REGION Network 43
   RUNG wire#powerrail
      Contact( "DB92".Static_1 )
      { S7_GenerateENO := "TRUE" } Move(in := 1, out1 => "DB46".Static_19)
      wire#w1
      Coil( "Tag_6" )
   END_RUNG
   RUNG wire#powerrail
      I_Contact( "DB92".Static_1 )
      { S7_GenerateENO := "TRUE" } Move(in := 2, out1 => "DB46".Static_19)
   END_RUNG wire#w1
   // the same network as SCL:
   // ENO of a box is taken as its EN; it also drops when the box reports an error
   IF "DB92".Static_1 THEN "DB46".Static_19 := 1; END_IF;
   IF NOT "DB92".Static_1 THEN "DB46".Static_19 := 2; END_IF;
   "Tag_6" := "DB92".Static_1 OR NOT "DB92".Static_1;
END_REGION

REGION Network 44
   RUNG wire#powerrail
      Contact( "DB92".Static_2 )
      { S7_GenerateENO := "TRUE" } Move(in := 1, out1 => "DB46".Static_20)
      wire#w1
      Coil( "Tag_6" )
   END_RUNG
   RUNG wire#powerrail
      I_Contact( "DB92".Static_2 )
      { S7_GenerateENO := "TRUE" } Move(in := 2, out1 => "DB46".Static_20)
   END_RUNG wire#w1
   // the same network as SCL:
   // ENO of a box is taken as its EN; it also drops when the box reports an error
   IF "DB92".Static_2 THEN "DB46".Static_20 := 1; END_IF;
   IF NOT "DB92".Static_2 THEN "DB46".Static_20 := 2; END_IF;
   "Tag_6" := "DB92".Static_2 OR NOT "DB92".Static_2;
END_REGION

REGION Network 45
   RUNG wire#powerrail
      Contact( "DB21".Static_52 )
      { S7_GenerateENO := "TRUE" } Move(in := 1, out1 => "DB46".Static_23)
      wire#w1
      Coil( "Tag_6" )
   END_RUNG
   RUNG wire#powerrail
      I_Contact( "DB21".Static_52 )
      { S7_GenerateENO := "TRUE" } Move(in := 2, out1 => "DB46".Static_23)
   END_RUNG wire#w1
   // the same network as SCL:
   // ENO of a box is taken as its EN; it also drops when the box reports an error
   IF "DB21".Static_52 THEN "DB46".Static_23 := 1; END_IF;
   IF NOT "DB21".Static_52 THEN "DB46".Static_23 := 2; END_IF;
   "Tag_6" := "DB21".Static_52 OR NOT "DB21".Static_52;
END_REGION

REGION Network 46
   RUNG wire#powerrail
      Contact( "DB21".Static_53 )
      { S7_GenerateENO := "TRUE" } Move(in := 1, out1 => "DB46".Static_24)
      wire#w1
      Coil( "Tag_6" )
   END_RUNG
   RUNG wire#powerrail
      I_Contact( "DB21".Static_53 )
      { S7_GenerateENO := "TRUE" } Move(in := 2, out1 => "DB46".Static_24)
   END_RUNG wire#w1
   // the same network as SCL:
   // ENO of a box is taken as its EN; it also drops when the box reports an error
   IF "DB21".Static_53 THEN "DB46".Static_24 := 1; END_IF;
   IF NOT "DB21".Static_53 THEN "DB46".Static_24 := 2; END_IF;
   "Tag_6" := "DB21".Static_53 OR NOT "DB21".Static_53;
END_REGION

REGION Network 47
   RUNG wire#powerrail
      Contact( "DB135".Static_18 )
      { S7_GenerateENO := "TRUE" } Move(in := 0, out1 => "DB135".Static_0)
      wire#w1
      Coil( "Tag_6" )
   END_RUNG
   RUNG wire#powerrail
      I_Contact( "DB135".Static_18 )
      Contact( "DB88".Static_12 )
      { S7_GenerateENO := "TRUE" } Move(in := 1, out1 => "DB135".Static_0)
   END_RUNG wire#w1
   RUNG wire#powerrail
      I_Contact( "DB135".Static_18 )
      I_Contact( "DB88".Static_12 )
      { S7_GenerateENO := "TRUE" } Move(in := 2, out1 => "DB135".Static_0)
   END_RUNG wire#w1
   // the same network as SCL:
   // ENO of a box is taken as its EN; it also drops when the box reports an error
   IF "DB135".Static_18 THEN "DB135".Static_0 := 0; END_IF;
   #_w1 := NOT "DB135".Static_18 AND "DB88".Static_12;
   IF #_w1 THEN "DB135".Static_0 := 1; END_IF;
   #_w2 := NOT "DB135".Static_18 AND NOT "DB88".Static_12;
   IF #_w2 THEN "DB135".Static_0 := 2; END_IF;
   "Tag_6" := "DB135".Static_18 OR #_w1 OR #_w2;
END_REGION

REGION Network 48
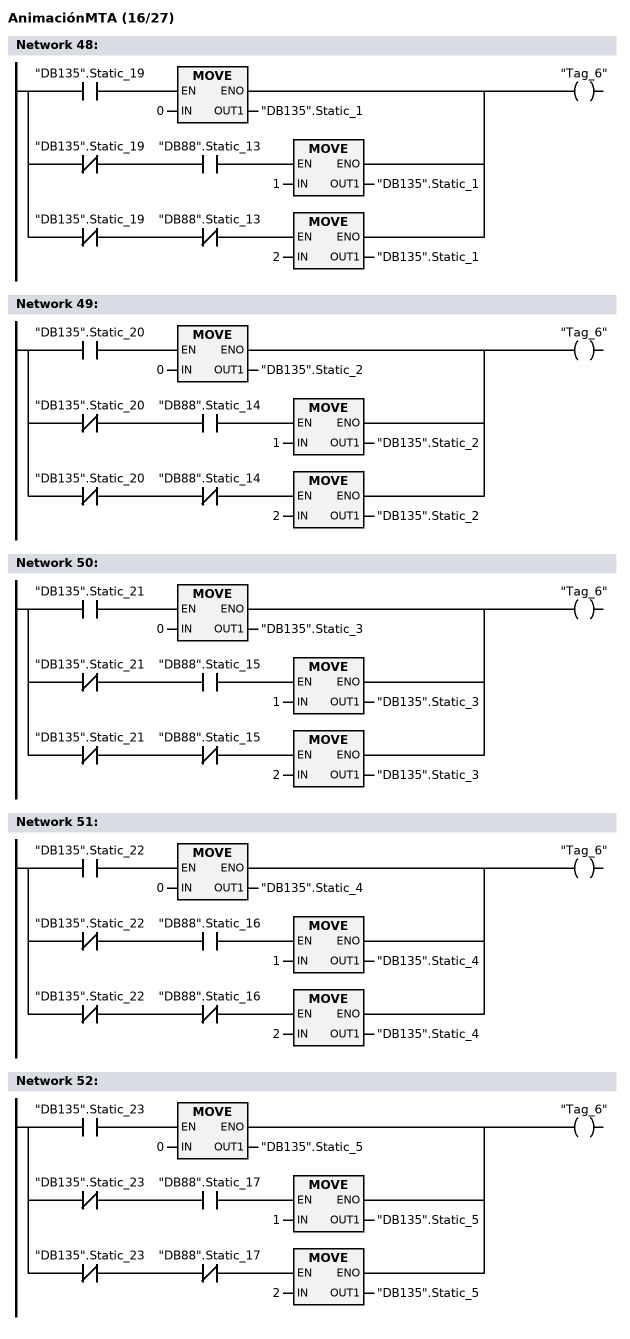
   RUNG wire#powerrail
      Contact( "DB135".Static_19 )
      { S7_GenerateENO := "TRUE" } Move(in := 0, out1 => "DB135".Static_1)
      wire#w1
      Coil( "Tag_6" )
   END_RUNG
   RUNG wire#powerrail
      I_Contact( "DB135".Static_19 )
      Contact( "DB88".Static_13 )
      { S7_GenerateENO := "TRUE" } Move(in := 1, out1 => "DB135".Static_1)
   END_RUNG wire#w1
   RUNG wire#powerrail
      I_Contact( "DB135".Static_19 )
      I_Contact( "DB88".Static_13 )
      { S7_GenerateENO := "TRUE" } Move(in := 2, out1 => "DB135".Static_1)
   END_RUNG wire#w1
   // the same network as SCL:
   // ENO of a box is taken as its EN; it also drops when the box reports an error
   IF "DB135".Static_19 THEN "DB135".Static_1 := 0; END_IF;
   #_w1 := NOT "DB135".Static_19 AND "DB88".Static_13;
   IF #_w1 THEN "DB135".Static_1 := 1; END_IF;
   #_w2 := NOT "DB135".Static_19 AND NOT "DB88".Static_13;
   IF #_w2 THEN "DB135".Static_1 := 2; END_IF;
   "Tag_6" := "DB135".Static_19 OR #_w1 OR #_w2;
END_REGION

REGION Network 49
   RUNG wire#powerrail
      Contact( "DB135".Static_20 )
      { S7_GenerateENO := "TRUE" } Move(in := 0, out1 => "DB135".Static_2)
      wire#w1
      Coil( "Tag_6" )
   END_RUNG
   RUNG wire#powerrail
      I_Contact( "DB135".Static_20 )
      Contact( "DB88".Static_14 )
      { S7_GenerateENO := "TRUE" } Move(in := 1, out1 => "DB135".Static_2)
   END_RUNG wire#w1
   RUNG wire#powerrail
      I_Contact( "DB135".Static_20 )
      I_Contact( "DB88".Static_14 )
      { S7_GenerateENO := "TRUE" } Move(in := 2, out1 => "DB135".Static_2)
   END_RUNG wire#w1
   // the same network as SCL:
   // ENO of a box is taken as its EN; it also drops when the box reports an error
   IF "DB135".Static_20 THEN "DB135".Static_2 := 0; END_IF;
   #_w1 := NOT "DB135".Static_20 AND "DB88".Static_14;
   IF #_w1 THEN "DB135".Static_2 := 1; END_IF;
   #_w2 := NOT "DB135".Static_20 AND NOT "DB88".Static_14;
   IF #_w2 THEN "DB135".Static_2 := 2; END_IF;
   "Tag_6" := "DB135".Static_20 OR #_w1 OR #_w2;
END_REGION

REGION Network 50
   RUNG wire#powerrail
      Contact( "DB135".Static_21 )
      { S7_GenerateENO := "TRUE" } Move(in := 0, out1 => "DB135".Static_3)
      wire#w1
      Coil( "Tag_6" )
   END_RUNG
   RUNG wire#powerrail
      I_Contact( "DB135".Static_21 )
      Contact( "DB88".Static_15 )
      { S7_GenerateENO := "TRUE" } Move(in := 1, out1 => "DB135".Static_3)
   END_RUNG wire#w1
   RUNG wire#powerrail
      I_Contact( "DB135".Static_21 )
      I_Contact( "DB88".Static_15 )
      { S7_GenerateENO := "TRUE" } Move(in := 2, out1 => "DB135".Static_3)
   END_RUNG wire#w1
   // the same network as SCL:
   // ENO of a box is taken as its EN; it also drops when the box reports an error
   IF "DB135".Static_21 THEN "DB135".Static_3 := 0; END_IF;
   #_w1 := NOT "DB135".Static_21 AND "DB88".Static_15;
   IF #_w1 THEN "DB135".Static_3 := 1; END_IF;
   #_w2 := NOT "DB135".Static_21 AND NOT "DB88".Static_15;
   IF #_w2 THEN "DB135".Static_3 := 2; END_IF;
   "Tag_6" := "DB135".Static_21 OR #_w1 OR #_w2;
END_REGION

REGION Network 51
   RUNG wire#powerrail
      Contact( "DB135".Static_22 )
      { S7_GenerateENO := "TRUE" } Move(in := 0, out1 => "DB135".Static_4)
      wire#w1
      Coil( "Tag_6" )
   END_RUNG
   RUNG wire#powerrail
      I_Contact( "DB135".Static_22 )
      Contact( "DB88".Static_16 )
      { S7_GenerateENO := "TRUE" } Move(in := 1, out1 => "DB135".Static_4)
   END_RUNG wire#w1
   RUNG wire#powerrail
      I_Contact( "DB135".Static_22 )
      I_Contact( "DB88".Static_16 )
      { S7_GenerateENO := "TRUE" } Move(in := 2, out1 => "DB135".Static_4)
   END_RUNG wire#w1
   // the same network as SCL:
   // ENO of a box is taken as its EN; it also drops when the box reports an error
   IF "DB135".Static_22 THEN "DB135".Static_4 := 0; END_IF;
   #_w1 := NOT "DB135".Static_22 AND "DB88".Static_16;
   IF #_w1 THEN "DB135".Static_4 := 1; END_IF;
   #_w2 := NOT "DB135".Static_22 AND NOT "DB88".Static_16;
   IF #_w2 THEN "DB135".Static_4 := 2; END_IF;
   "Tag_6" := "DB135".Static_22 OR #_w1 OR #_w2;
END_REGION

REGION Network 52
   RUNG wire#powerrail
      Contact( "DB135".Static_23 )
      { S7_GenerateENO := "TRUE" } Move(in := 0, out1 => "DB135".Static_5)
      wire#w1
      Coil( "Tag_6" )
   END_RUNG
   RUNG wire#powerrail
      I_Contact( "DB135".Static_23 )
      Contact( "DB88".Static_17 )
      { S7_GenerateENO := "TRUE" } Move(in := 1, out1 => "DB135".Static_5)
   END_RUNG wire#w1
   RUNG wire#powerrail
      I_Contact( "DB135".Static_23 )
      I_Contact( "DB88".Static_17 )
      { S7_GenerateENO := "TRUE" } Move(in := 2, out1 => "DB135".Static_5)
   END_RUNG wire#w1
   // the same network as SCL:
   // ENO of a box is taken as its EN; it also drops when the box reports an error
   IF "DB135".Static_23 THEN "DB135".Static_5 := 0; END_IF;
   #_w1 := NOT "DB135".Static_23 AND "DB88".Static_17;
   IF #_w1 THEN "DB135".Static_5 := 1; END_IF;
   #_w2 := NOT "DB135".Static_23 AND NOT "DB88".Static_17;
   IF #_w2 THEN "DB135".Static_5 := 2; END_IF;
   "Tag_6" := "DB135".Static_23 OR #_w1 OR #_w2;
END_REGION

REGION Network 53
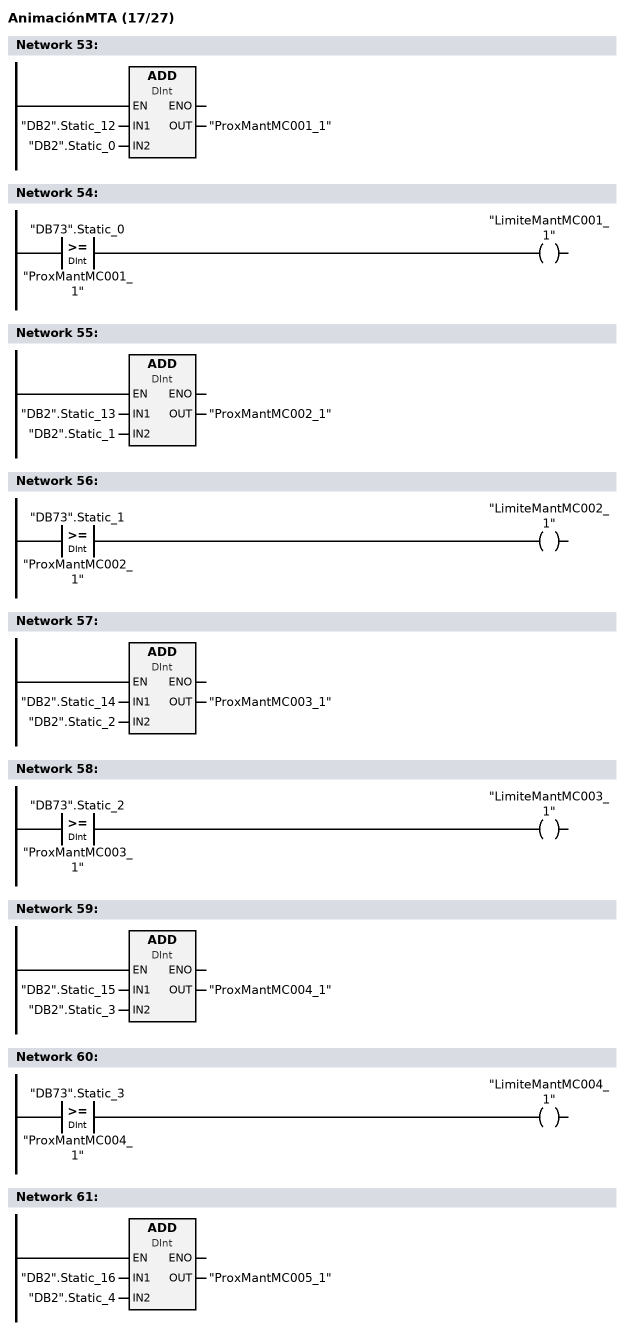
   RUNG wire#powerrail
      { S7_Templates := "SrcType := DInt"; S7_GenerateENO := "TRUE" } Add(in1 := "DB2".Static_12, in2 := "DB2".Static_0, out => "ProxMantMC001_1")
   END_RUNG
   // the same network as SCL:
   "ProxMantMC001_1" := "DB2".Static_12 + "DB2".Static_0;
END_REGION

REGION Network 54
   RUNG wire#powerrail
      { S7_Templates := "SrcType := DInt" } GE_Contact(in1 := "DB73".Static_0, in2 := "ProxMantMC001_1")
      Coil( "LimiteMantMC001_1" )
   END_RUNG
   // the same network as SCL:
   "LimiteMantMC001_1" := "DB73".Static_0 >= "ProxMantMC001_1";
END_REGION

REGION Network 55
   RUNG wire#powerrail
      { S7_Templates := "SrcType := DInt"; S7_GenerateENO := "TRUE" } Add(in1 := "DB2".Static_13, in2 := "DB2".Static_1, out => "ProxMantMC002_1")
   END_RUNG
   // the same network as SCL:
   "ProxMantMC002_1" := "DB2".Static_13 + "DB2".Static_1;
END_REGION

REGION Network 56
   RUNG wire#powerrail
      { S7_Templates := "SrcType := DInt" } GE_Contact(in1 := "DB73".Static_1, in2 := "ProxMantMC002_1")
      Coil( "LimiteMantMC002_1" )
   END_RUNG
   // the same network as SCL:
   "LimiteMantMC002_1" := "DB73".Static_1 >= "ProxMantMC002_1";
END_REGION

REGION Network 57
   RUNG wire#powerrail
      { S7_Templates := "SrcType := DInt"; S7_GenerateENO := "TRUE" } Add(in1 := "DB2".Static_14, in2 := "DB2".Static_2, out => "ProxMantMC003_1")
   END_RUNG
   // the same network as SCL:
   "ProxMantMC003_1" := "DB2".Static_14 + "DB2".Static_2;
END_REGION

REGION Network 58
   RUNG wire#powerrail
      { S7_Templates := "SrcType := DInt" } GE_Contact(in1 := "DB73".Static_2, in2 := "ProxMantMC003_1")
      Coil( "LimiteMantMC003_1" )
   END_RUNG
   // the same network as SCL:
   "LimiteMantMC003_1" := "DB73".Static_2 >= "ProxMantMC003_1";
END_REGION

REGION Network 59
   RUNG wire#powerrail
      { S7_Templates := "SrcType := DInt"; S7_GenerateENO := "TRUE" } Add(in1 := "DB2".Static_15, in2 := "DB2".Static_3, out => "ProxMantMC004_1")
   END_RUNG
   // the same network as SCL:
   "ProxMantMC004_1" := "DB2".Static_15 + "DB2".Static_3;
END_REGION

REGION Network 60
   RUNG wire#powerrail
      { S7_Templates := "SrcType := DInt" } GE_Contact(in1 := "DB73".Static_3, in2 := "ProxMantMC004_1")
      Coil( "LimiteMantMC004_1" )
   END_RUNG
   // the same network as SCL:
   "LimiteMantMC004_1" := "DB73".Static_3 >= "ProxMantMC004_1";
END_REGION

REGION Network 61
   RUNG wire#powerrail
      { S7_Templates := "SrcType := DInt"; S7_GenerateENO := "TRUE" } Add(in1 := "DB2".Static_16, in2 := "DB2".Static_4, out => "ProxMantMC005_1")
   END_RUNG
   // the same network as SCL:
   "ProxMantMC005_1" := "DB2".Static_16 + "DB2".Static_4;
END_REGION

REGION Network 62
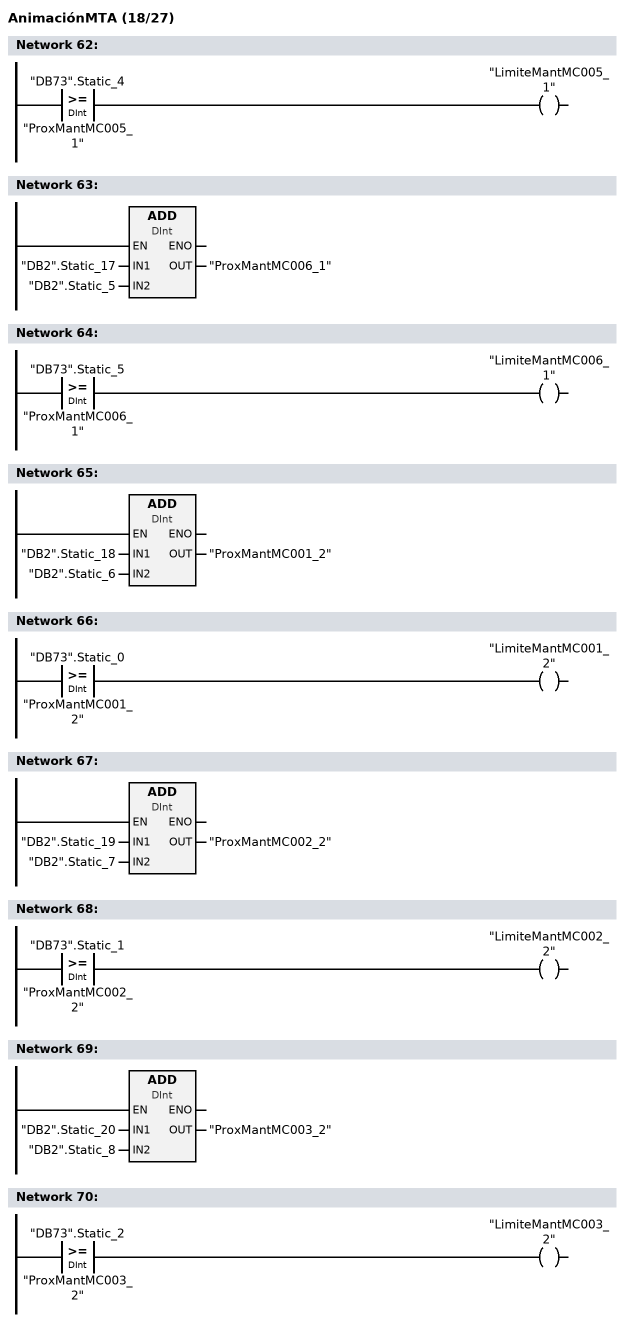
   RUNG wire#powerrail
      { S7_Templates := "SrcType := DInt" } GE_Contact(in1 := "DB73".Static_4, in2 := "ProxMantMC005_1")
      Coil( "LimiteMantMC005_1" )
   END_RUNG
   // the same network as SCL:
   "LimiteMantMC005_1" := "DB73".Static_4 >= "ProxMantMC005_1";
END_REGION

REGION Network 63
   RUNG wire#powerrail
      { S7_Templates := "SrcType := DInt"; S7_GenerateENO := "TRUE" } Add(in1 := "DB2".Static_17, in2 := "DB2".Static_5, out => "ProxMantMC006_1")
   END_RUNG
   // the same network as SCL:
   "ProxMantMC006_1" := "DB2".Static_17 + "DB2".Static_5;
END_REGION

REGION Network 64
   RUNG wire#powerrail
      { S7_Templates := "SrcType := DInt" } GE_Contact(in1 := "DB73".Static_5, in2 := "ProxMantMC006_1")
      Coil( "LimiteMantMC006_1" )
   END_RUNG
   // the same network as SCL:
   "LimiteMantMC006_1" := "DB73".Static_5 >= "ProxMantMC006_1";
END_REGION

REGION Network 65
   RUNG wire#powerrail
      { S7_Templates := "SrcType := DInt"; S7_GenerateENO := "TRUE" } Add(in1 := "DB2".Static_18, in2 := "DB2".Static_6, out => "ProxMantMC001_2")
   END_RUNG
   // the same network as SCL:
   "ProxMantMC001_2" := "DB2".Static_18 + "DB2".Static_6;
END_REGION

REGION Network 66
   RUNG wire#powerrail
      { S7_Templates := "SrcType := DInt" } GE_Contact(in1 := "DB73".Static_0, in2 := "ProxMantMC001_2")
      Coil( "LimiteMantMC001_2" )
   END_RUNG
   // the same network as SCL:
   "LimiteMantMC001_2" := "DB73".Static_0 >= "ProxMantMC001_2";
END_REGION

REGION Network 67
   RUNG wire#powerrail
      { S7_Templates := "SrcType := DInt"; S7_GenerateENO := "TRUE" } Add(in1 := "DB2".Static_19, in2 := "DB2".Static_7, out => "ProxMantMC002_2")
   END_RUNG
   // the same network as SCL:
   "ProxMantMC002_2" := "DB2".Static_19 + "DB2".Static_7;
END_REGION

REGION Network 68
   RUNG wire#powerrail
      { S7_Templates := "SrcType := DInt" } GE_Contact(in1 := "DB73".Static_1, in2 := "ProxMantMC002_2")
      Coil( "LimiteMantMC002_2" )
   END_RUNG
   // the same network as SCL:
   "LimiteMantMC002_2" := "DB73".Static_1 >= "ProxMantMC002_2";
END_REGION

REGION Network 69
   RUNG wire#powerrail
      { S7_Templates := "SrcType := DInt"; S7_GenerateENO := "TRUE" } Add(in1 := "DB2".Static_20, in2 := "DB2".Static_8, out => "ProxMantMC003_2")
   END_RUNG
   // the same network as SCL:
   "ProxMantMC003_2" := "DB2".Static_20 + "DB2".Static_8;
END_REGION

REGION Network 70
   RUNG wire#powerrail
      { S7_Templates := "SrcType := DInt" } GE_Contact(in1 := "DB73".Static_2, in2 := "ProxMantMC003_2")
      Coil( "LimiteMantMC003_2" )
   END_RUNG
   // the same network as SCL:
   "LimiteMantMC003_2" := "DB73".Static_2 >= "ProxMantMC003_2";
END_REGION

REGION Network 71
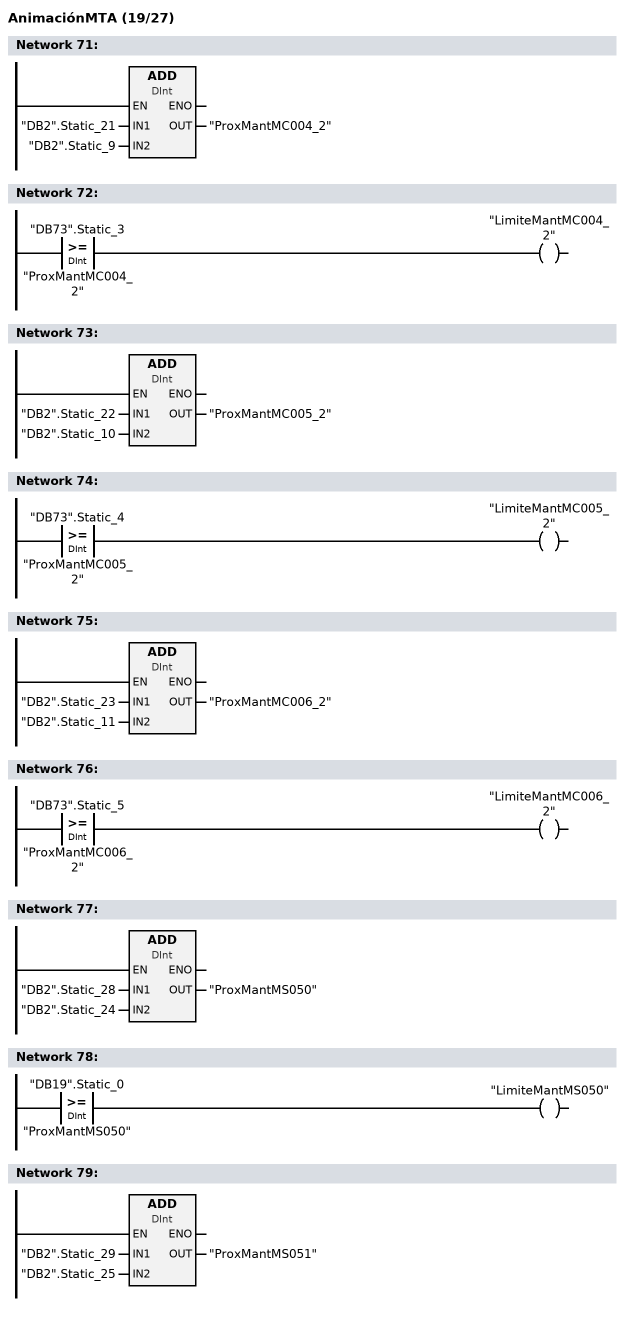
   RUNG wire#powerrail
      { S7_Templates := "SrcType := DInt"; S7_GenerateENO := "TRUE" } Add(in1 := "DB2".Static_21, in2 := "DB2".Static_9, out => "ProxMantMC004_2")
   END_RUNG
   // the same network as SCL:
   "ProxMantMC004_2" := "DB2".Static_21 + "DB2".Static_9;
END_REGION

REGION Network 72
   RUNG wire#powerrail
      { S7_Templates := "SrcType := DInt" } GE_Contact(in1 := "DB73".Static_3, in2 := "ProxMantMC004_2")
      Coil( "LimiteMantMC004_2" )
   END_RUNG
   // the same network as SCL:
   "LimiteMantMC004_2" := "DB73".Static_3 >= "ProxMantMC004_2";
END_REGION

REGION Network 73
   RUNG wire#powerrail
      { S7_Templates := "SrcType := DInt"; S7_GenerateENO := "TRUE" } Add(in1 := "DB2".Static_22, in2 := "DB2".Static_10, out => "ProxMantMC005_2")
   END_RUNG
   // the same network as SCL:
   "ProxMantMC005_2" := "DB2".Static_22 + "DB2".Static_10;
END_REGION

REGION Network 74
   RUNG wire#powerrail
      { S7_Templates := "SrcType := DInt" } GE_Contact(in1 := "DB73".Static_4, in2 := "ProxMantMC005_2")
      Coil( "LimiteMantMC005_2" )
   END_RUNG
   // the same network as SCL:
   "LimiteMantMC005_2" := "DB73".Static_4 >= "ProxMantMC005_2";
END_REGION

REGION Network 75
   RUNG wire#powerrail
      { S7_Templates := "SrcType := DInt"; S7_GenerateENO := "TRUE" } Add(in1 := "DB2".Static_23, in2 := "DB2".Static_11, out => "ProxMantMC006_2")
   END_RUNG
   // the same network as SCL:
   "ProxMantMC006_2" := "DB2".Static_23 + "DB2".Static_11;
END_REGION

REGION Network 76
   RUNG wire#powerrail
      { S7_Templates := "SrcType := DInt" } GE_Contact(in1 := "DB73".Static_5, in2 := "ProxMantMC006_2")
      Coil( "LimiteMantMC006_2" )
   END_RUNG
   // the same network as SCL:
   "LimiteMantMC006_2" := "DB73".Static_5 >= "ProxMantMC006_2";
END_REGION

REGION Network 77
   RUNG wire#powerrail
      { S7_Templates := "SrcType := DInt"; S7_GenerateENO := "TRUE" } Add(in1 := "DB2".Static_28, in2 := "DB2".Static_24, out => "ProxMantMS050")
   END_RUNG
   // the same network as SCL:
   "ProxMantMS050" := "DB2".Static_28 + "DB2".Static_24;
END_REGION

REGION Network 78
   RUNG wire#powerrail
      { S7_Templates := "SrcType := DInt" } GE_Contact(in1 := "DB19".Static_0, in2 := "ProxMantMS050")
      Coil( "LimiteMantMS050" )
   END_RUNG
   // the same network as SCL:
   "LimiteMantMS050" := "DB19".Static_0 >= "ProxMantMS050";
END_REGION

REGION Network 79
   RUNG wire#powerrail
      { S7_Templates := "SrcType := DInt"; S7_GenerateENO := "TRUE" } Add(in1 := "DB2".Static_29, in2 := "DB2".Static_25, out => "ProxMantMS051")
   END_RUNG
   // the same network as SCL:
   "ProxMantMS051" := "DB2".Static_29 + "DB2".Static_25;
END_REGION

REGION Network 80
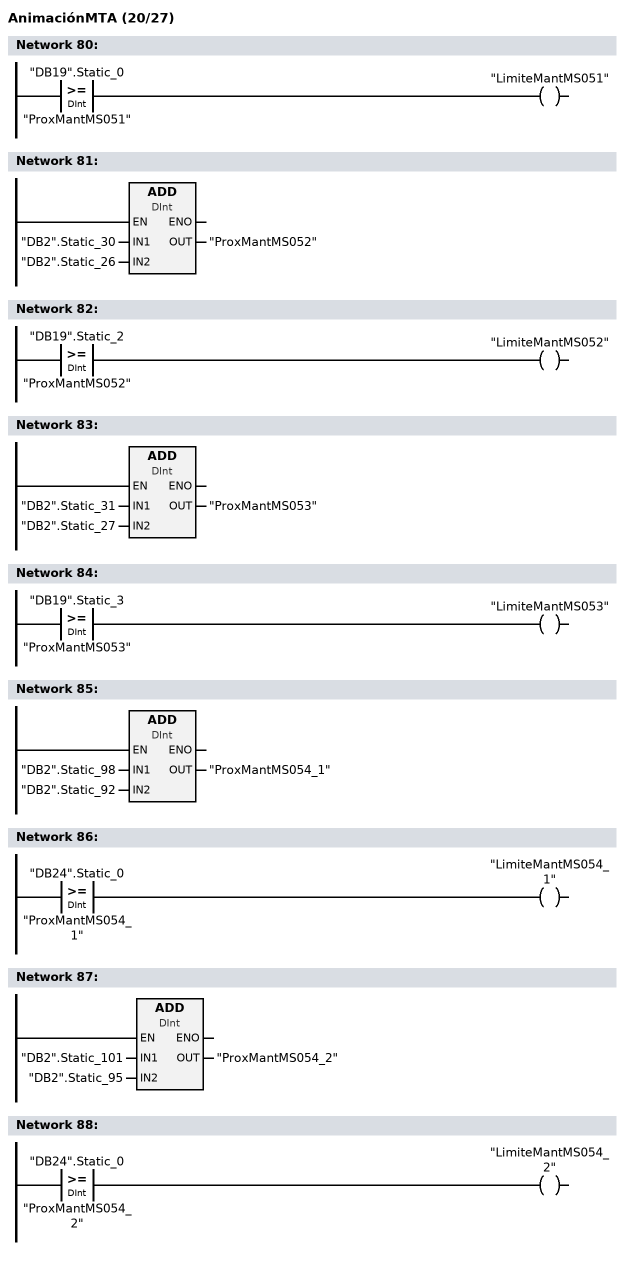
   RUNG wire#powerrail
      { S7_Templates := "SrcType := DInt" } GE_Contact(in1 := "DB19".Static_0, in2 := "ProxMantMS051")
      Coil( "LimiteMantMS051" )
   END_RUNG
   // the same network as SCL:
   "LimiteMantMS051" := "DB19".Static_0 >= "ProxMantMS051";
END_REGION

REGION Network 81
   RUNG wire#powerrail
      { S7_Templates := "SrcType := DInt"; S7_GenerateENO := "TRUE" } Add(in1 := "DB2".Static_30, in2 := "DB2".Static_26, out => "ProxMantMS052")
   END_RUNG
   // the same network as SCL:
   "ProxMantMS052" := "DB2".Static_30 + "DB2".Static_26;
END_REGION

REGION Network 82
   RUNG wire#powerrail
      { S7_Templates := "SrcType := DInt" } GE_Contact(in1 := "DB19".Static_2, in2 := "ProxMantMS052")
      Coil( "LimiteMantMS052" )
   END_RUNG
   // the same network as SCL:
   "LimiteMantMS052" := "DB19".Static_2 >= "ProxMantMS052";
END_REGION

REGION Network 83
   RUNG wire#powerrail
      { S7_Templates := "SrcType := DInt"; S7_GenerateENO := "TRUE" } Add(in1 := "DB2".Static_31, in2 := "DB2".Static_27, out => "ProxMantMS053")
   END_RUNG
   // the same network as SCL:
   "ProxMantMS053" := "DB2".Static_31 + "DB2".Static_27;
END_REGION

REGION Network 84
   RUNG wire#powerrail
      { S7_Templates := "SrcType := DInt" } GE_Contact(in1 := "DB19".Static_3, in2 := "ProxMantMS053")
      Coil( "LimiteMantMS053" )
   END_RUNG
   // the same network as SCL:
   "LimiteMantMS053" := "DB19".Static_3 >= "ProxMantMS053";
END_REGION

REGION Network 85
   RUNG wire#powerrail
      { S7_Templates := "SrcType := DInt"; S7_GenerateENO := "TRUE" } Add(in1 := "DB2".Static_98, in2 := "DB2".Static_92, out => "ProxMantMS054_1")
   END_RUNG
   // the same network as SCL:
   "ProxMantMS054_1" := "DB2".Static_98 + "DB2".Static_92;
END_REGION

REGION Network 86
   RUNG wire#powerrail
      { S7_Templates := "SrcType := DInt" } GE_Contact(in1 := "DB24".Static_0, in2 := "ProxMantMS054_1")
      Coil( "LimiteMantMS054_1" )
   END_RUNG
   // the same network as SCL:
   "LimiteMantMS054_1" := "DB24".Static_0 >= "ProxMantMS054_1";
END_REGION

REGION Network 87
   RUNG wire#powerrail
      { S7_Templates := "SrcType := DInt"; S7_GenerateENO := "TRUE" } Add(in1 := "DB2".Static_101, in2 := "DB2".Static_95, out => "ProxMantMS054_2")
   END_RUNG
   // the same network as SCL:
   "ProxMantMS054_2" := "DB2".Static_101 + "DB2".Static_95;
END_REGION

REGION Network 88
   RUNG wire#powerrail
      { S7_Templates := "SrcType := DInt" } GE_Contact(in1 := "DB24".Static_0, in2 := "ProxMantMS054_2")
      Coil( "LimiteMantMS054_2" )
   END_RUNG
   // the same network as SCL:
   "LimiteMantMS054_2" := "DB24".Static_0 >= "ProxMantMS054_2";
END_REGION

REGION Network 89
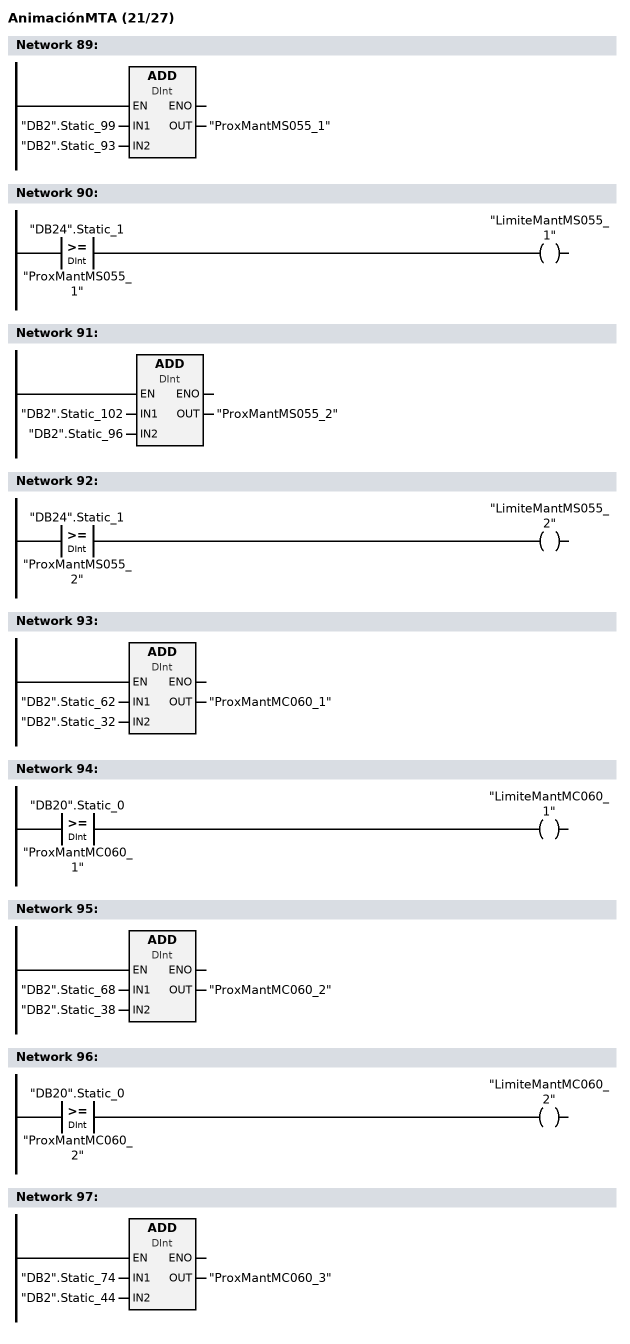
   RUNG wire#powerrail
      { S7_Templates := "SrcType := DInt"; S7_GenerateENO := "TRUE" } Add(in1 := "DB2".Static_99, in2 := "DB2".Static_93, out => "ProxMantMS055_1")
   END_RUNG
   // the same network as SCL:
   "ProxMantMS055_1" := "DB2".Static_99 + "DB2".Static_93;
END_REGION

REGION Network 90
   RUNG wire#powerrail
      { S7_Templates := "SrcType := DInt" } GE_Contact(in1 := "DB24".Static_1, in2 := "ProxMantMS055_1")
      Coil( "LimiteMantMS055_1" )
   END_RUNG
   // the same network as SCL:
   "LimiteMantMS055_1" := "DB24".Static_1 >= "ProxMantMS055_1";
END_REGION

REGION Network 91
   RUNG wire#powerrail
      { S7_Templates := "SrcType := DInt"; S7_GenerateENO := "TRUE" } Add(in1 := "DB2".Static_102, in2 := "DB2".Static_96, out => "ProxMantMS055_2")
   END_RUNG
   // the same network as SCL:
   "ProxMantMS055_2" := "DB2".Static_102 + "DB2".Static_96;
END_REGION

REGION Network 92
   RUNG wire#powerrail
      { S7_Templates := "SrcType := DInt" } GE_Contact(in1 := "DB24".Static_1, in2 := "ProxMantMS055_2")
      Coil( "LimiteMantMS055_2" )
   END_RUNG
   // the same network as SCL:
   "LimiteMantMS055_2" := "DB24".Static_1 >= "ProxMantMS055_2";
END_REGION

REGION Network 93
   RUNG wire#powerrail
      { S7_Templates := "SrcType := DInt"; S7_GenerateENO := "TRUE" } Add(in1 := "DB2".Static_62, in2 := "DB2".Static_32, out => "ProxMantMC060_1")
   END_RUNG
   // the same network as SCL:
   "ProxMantMC060_1" := "DB2".Static_62 + "DB2".Static_32;
END_REGION

REGION Network 94
   RUNG wire#powerrail
      { S7_Templates := "SrcType := DInt" } GE_Contact(in1 := "DB20".Static_0, in2 := "ProxMantMC060_1")
      Coil( "LimiteMantMC060_1" )
   END_RUNG
   // the same network as SCL:
   "LimiteMantMC060_1" := "DB20".Static_0 >= "ProxMantMC060_1";
END_REGION

REGION Network 95
   RUNG wire#powerrail
      { S7_Templates := "SrcType := DInt"; S7_GenerateENO := "TRUE" } Add(in1 := "DB2".Static_68, in2 := "DB2".Static_38, out => "ProxMantMC060_2")
   END_RUNG
   // the same network as SCL:
   "ProxMantMC060_2" := "DB2".Static_68 + "DB2".Static_38;
END_REGION

REGION Network 96
   RUNG wire#powerrail
      { S7_Templates := "SrcType := DInt" } GE_Contact(in1 := "DB20".Static_0, in2 := "ProxMantMC060_2")
      Coil( "LimiteMantMC060_2" )
   END_RUNG
   // the same network as SCL:
   "LimiteMantMC060_2" := "DB20".Static_0 >= "ProxMantMC060_2";
END_REGION

REGION Network 97
   RUNG wire#powerrail
      { S7_Templates := "SrcType := DInt"; S7_GenerateENO := "TRUE" } Add(in1 := "DB2".Static_74, in2 := "DB2".Static_44, out => "ProxMantMC060_3")
   END_RUNG
   // the same network as SCL:
   "ProxMantMC060_3" := "DB2".Static_74 + "DB2".Static_44;
END_REGION

REGION Network 98
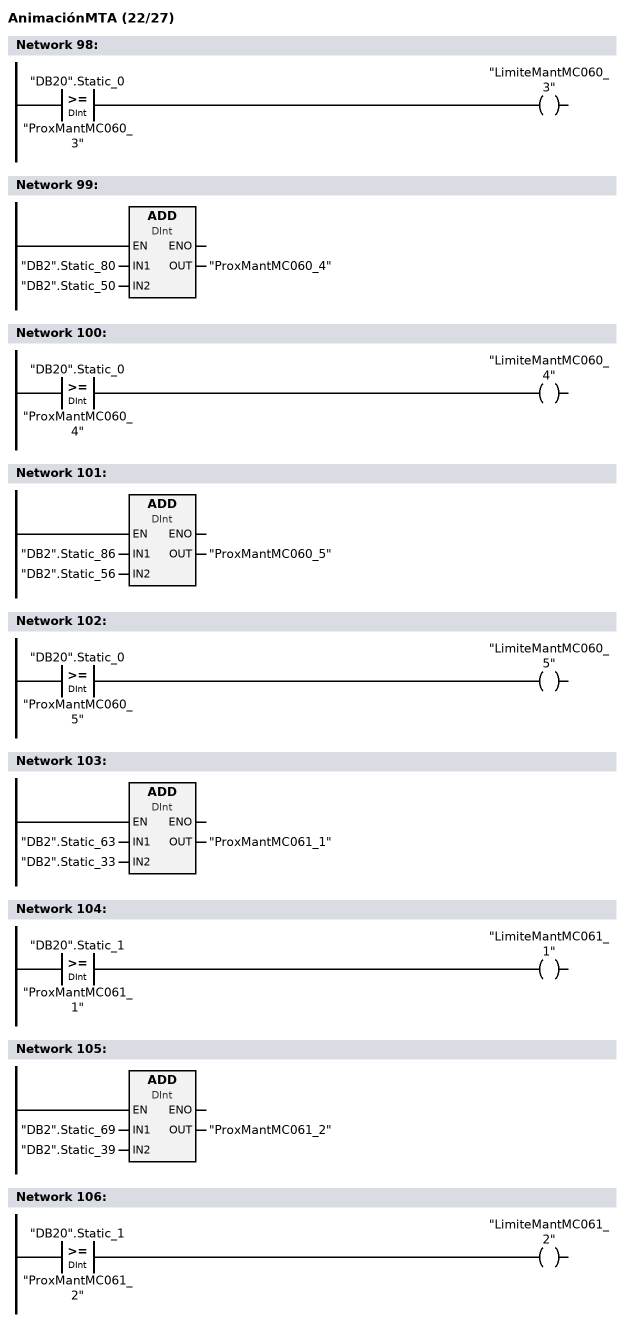
   RUNG wire#powerrail
      { S7_Templates := "SrcType := DInt" } GE_Contact(in1 := "DB20".Static_0, in2 := "ProxMantMC060_3")
      Coil( "LimiteMantMC060_3" )
   END_RUNG
   // the same network as SCL:
   "LimiteMantMC060_3" := "DB20".Static_0 >= "ProxMantMC060_3";
END_REGION

REGION Network 99
   RUNG wire#powerrail
      { S7_Templates := "SrcType := DInt"; S7_GenerateENO := "TRUE" } Add(in1 := "DB2".Static_80, in2 := "DB2".Static_50, out => "ProxMantMC060_4")
   END_RUNG
   // the same network as SCL:
   "ProxMantMC060_4" := "DB2".Static_80 + "DB2".Static_50;
END_REGION

REGION Network 100
   RUNG wire#powerrail
      { S7_Templates := "SrcType := DInt" } GE_Contact(in1 := "DB20".Static_0, in2 := "ProxMantMC060_4")
      Coil( "LimiteMantMC060_4" )
   END_RUNG
   // the same network as SCL:
   "LimiteMantMC060_4" := "DB20".Static_0 >= "ProxMantMC060_4";
END_REGION

REGION Network 101
   RUNG wire#powerrail
      { S7_Templates := "SrcType := DInt"; S7_GenerateENO := "TRUE" } Add(in1 := "DB2".Static_86, in2 := "DB2".Static_56, out => "ProxMantMC060_5")
   END_RUNG
   // the same network as SCL:
   "ProxMantMC060_5" := "DB2".Static_86 + "DB2".Static_56;
END_REGION

REGION Network 102
   RUNG wire#powerrail
      { S7_Templates := "SrcType := DInt" } GE_Contact(in1 := "DB20".Static_0, in2 := "ProxMantMC060_5")
      Coil( "LimiteMantMC060_5" )
   END_RUNG
   // the same network as SCL:
   "LimiteMantMC060_5" := "DB20".Static_0 >= "ProxMantMC060_5";
END_REGION

REGION Network 103
   RUNG wire#powerrail
      { S7_Templates := "SrcType := DInt"; S7_GenerateENO := "TRUE" } Add(in1 := "DB2".Static_63, in2 := "DB2".Static_33, out => "ProxMantMC061_1")
   END_RUNG
   // the same network as SCL:
   "ProxMantMC061_1" := "DB2".Static_63 + "DB2".Static_33;
END_REGION

REGION Network 104
   RUNG wire#powerrail
      { S7_Templates := "SrcType := DInt" } GE_Contact(in1 := "DB20".Static_1, in2 := "ProxMantMC061_1")
      Coil( "LimiteMantMC061_1" )
   END_RUNG
   // the same network as SCL:
   "LimiteMantMC061_1" := "DB20".Static_1 >= "ProxMantMC061_1";
END_REGION

REGION Network 105
   RUNG wire#powerrail
      { S7_Templates := "SrcType := DInt"; S7_GenerateENO := "TRUE" } Add(in1 := "DB2".Static_69, in2 := "DB2".Static_39, out => "ProxMantMC061_2")
   END_RUNG
   // the same network as SCL:
   "ProxMantMC061_2" := "DB2".Static_69 + "DB2".Static_39;
END_REGION

REGION Network 106
   RUNG wire#powerrail
      { S7_Templates := "SrcType := DInt" } GE_Contact(in1 := "DB20".Static_1, in2 := "ProxMantMC061_2")
      Coil( "LimiteMantMC061_2" )
   END_RUNG
   // the same network as SCL:
   "LimiteMantMC061_2" := "DB20".Static_1 >= "ProxMantMC061_2";
END_REGION

REGION Network 107
